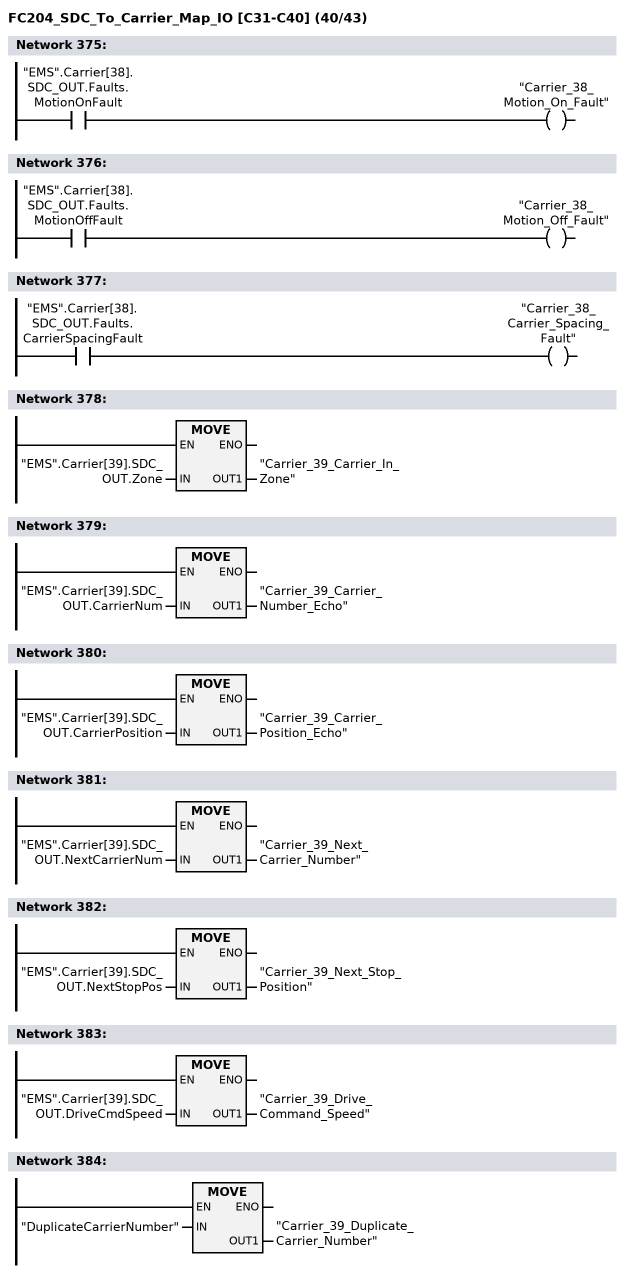
   RUNG wire#powerrail
      Contact( "EMS".Carrier[38].SDC_OUT.Faults.MotionOnFault )
      Coil( "Carrier_38_Motion_On_Fault" )
   END_RUNG
   // the same network as SCL:
   "Carrier_38_Motion_On_Fault" := "EMS".Carrier[38].SDC_OUT.Faults.MotionOnFault;
END_REGION

REGION Network 376
   RUNG wire#powerrail
      Contact( "EMS".Carrier[38].SDC_OUT.Faults.MotionOffFault )
      Coil( "Carrier_38_Motion_Off_Fault" )
   END_RUNG
   // the same network as SCL:
   "Carrier_38_Motion_Off_Fault" := "EMS".Carrier[38].SDC_OUT.Faults.MotionOffFault;
END_REGION

REGION Network 377
   RUNG wire#powerrail
      Contact( "EMS".Carrier[38].SDC_OUT.Faults.CarrierSpacingFault )
      Coil( "Carrier_38_Carrier_Spacing_Fault" )
   END_RUNG
   // the same network as SCL:
   "Carrier_38_Carrier_Spacing_Fault" := "EMS".Carrier[38].SDC_OUT.Faults.CarrierSpacingFault;
END_REGION

REGION Network 378
   RUNG wire#powerrail
      Move(in := "EMS".Carrier[39].SDC_OUT.Zone, out1 => "Carrier_39_Carrier_In_Zone")
   END_RUNG
   // the same network as SCL:
   "Carrier_39_Carrier_In_Zone" := "EMS".Carrier[39].SDC_OUT.Zone;
END_REGION

REGION Network 379
   RUNG wire#powerrail
      Move(in := "EMS".Carrier[39].SDC_OUT.CarrierNum, out1 => "Carrier_39_Carrier_Number_Echo")
   END_RUNG
   // the same network as SCL:
   "Carrier_39_Carrier_Number_Echo" := "EMS".Carrier[39].SDC_OUT.CarrierNum;
END_REGION

REGION Network 380
   RUNG wire#powerrail
      Move(in := "EMS".Carrier[39].SDC_OUT.CarrierPosition, out1 => "Carrier_39_Carrier_Position_Echo")
   END_RUNG
   // the same network as SCL:
   "Carrier_39_Carrier_Position_Echo" := "EMS".Carrier[39].SDC_OUT.CarrierPosition;
END_REGION

REGION Network 381
   RUNG wire#powerrail
      Move(in := "EMS".Carrier[39].SDC_OUT.NextCarrierNum, out1 => "Carrier_39_Next_Carrier_Number")
   END_RUNG
   // the same network as SCL:
   "Carrier_39_Next_Carrier_Number" := "EMS".Carrier[39].SDC_OUT.NextCarrierNum;
END_REGION

REGION Network 382
   RUNG wire#powerrail
      Move(in := "EMS".Carrier[39].SDC_OUT.NextStopPos, out1 => "Carrier_39_Next_Stop_Position")
   END_RUNG
   // the same network as SCL:
   "Carrier_39_Next_Stop_Position" := "EMS".Carrier[39].SDC_OUT.NextStopPos;
END_REGION

REGION Network 383
   RUNG wire#powerrail
      Move(in := "EMS".Carrier[39].SDC_OUT.DriveCmdSpeed, out1 => "Carrier_39_Drive_Command_Speed")
   END_RUNG
   // the same network as SCL:
   "Carrier_39_Drive_Command_Speed" := "EMS".Carrier[39].SDC_OUT.DriveCmdSpeed;
END_REGION

REGION Network 384
   RUNG wire#powerrail
      Move(in := "DuplicateCarrierNumber", out1 => "Carrier_39_Duplicate_Carrier_Number")
   END_RUNG
   // the same network as SCL:
   "Carrier_39_Duplicate_Carrier_Number" := "DuplicateCarrierNumber";
END_REGION

REGION Network 385
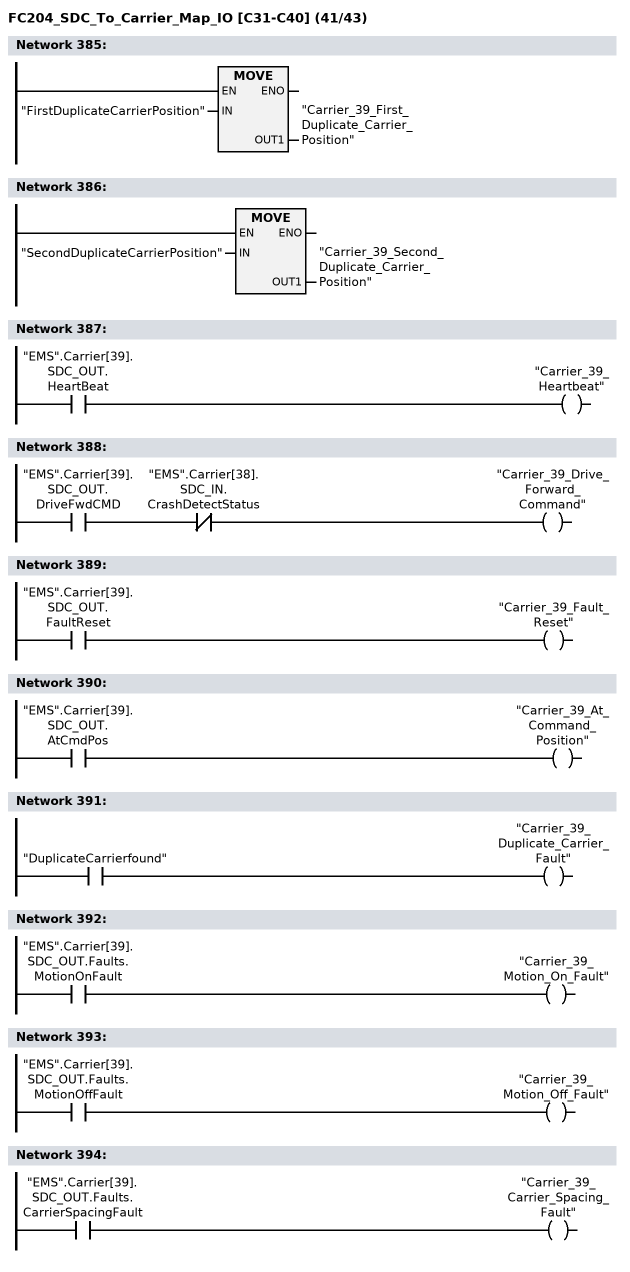
   RUNG wire#powerrail
      Move(in := "FirstDuplicateCarrierPosition", out1 => "Carrier_39_First_Duplicate_Carrier_Position")
   END_RUNG
   // the same network as SCL:
   "Carrier_39_First_Duplicate_Carrier_Position" := "FirstDuplicateCarrierPosition";
END_REGION

REGION Network 386
   RUNG wire#powerrail
      Move(in := "SecondDuplicateCarrierPosition", out1 => "Carrier_39_Second_Duplicate_Carrier_Position")
   END_RUNG
   // the same network as SCL:
   "Carrier_39_Second_Duplicate_Carrier_Position" := "SecondDuplicateCarrierPosition";
END_REGION

REGION Network 387
   RUNG wire#powerrail
      Contact( "EMS".Carrier[39].SDC_OUT.HeartBeat )
      Coil( "Carrier_39_Heartbeat" )
   END_RUNG
   // the same network as SCL:
   "Carrier_39_Heartbeat" := "EMS".Carrier[39].SDC_OUT.HeartBeat;
END_REGION

REGION Network 388
   RUNG wire#powerrail
      Contact( "EMS".Carrier[39].SDC_OUT.DriveFwdCMD )
      I_Contact( "EMS".Carrier[38].SDC_IN.CrashDetectStatus )
      Coil( "Carrier_39_Drive_Forward_Command" )
   END_RUNG
   // the same network as SCL:
   "Carrier_39_Drive_Forward_Command" := "EMS".Carrier[39].SDC_OUT.DriveFwdCMD AND NOT "EMS".Carrier[38].SDC_IN.CrashDetectStatus;
END_REGION

REGION Network 389
   RUNG wire#powerrail
      Contact( "EMS".Carrier[39].SDC_OUT.FaultReset )
      Coil( "Carrier_39_Fault_Reset" )
   END_RUNG
   // the same network as SCL:
   "Carrier_39_Fault_Reset" := "EMS".Carrier[39].SDC_OUT.FaultReset;
END_REGION

REGION Network 390
   RUNG wire#powerrail
      Contact( "EMS".Carrier[39].SDC_OUT.AtCmdPos )
      Coil( "Carrier_39_At_Command_Position" )
   END_RUNG
   // the same network as SCL:
   "Carrier_39_At_Command_Position" := "EMS".Carrier[39].SDC_OUT.AtCmdPos;
END_REGION

REGION Network 391
   RUNG wire#powerrail
      Contact( "DuplicateCarrierfound" )
      Coil( "Carrier_39_Duplicate_Carrier_Fault" )
   END_RUNG
   // the same network as SCL:
   "Carrier_39_Duplicate_Carrier_Fault" := "DuplicateCarrierfound";
END_REGION

REGION Network 392
   RUNG wire#powerrail
      Contact( "EMS".Carrier[39].SDC_OUT.Faults.MotionOnFault )
      Coil( "Carrier_39_Motion_On_Fault" )
   END_RUNG
   // the same network as SCL:
   "Carrier_39_Motion_On_Fault" := "EMS".Carrier[39].SDC_OUT.Faults.MotionOnFault;
END_REGION

REGION Network 393
   RUNG wire#powerrail
      Contact( "EMS".Carrier[39].SDC_OUT.Faults.MotionOffFault )
      Coil( "Carrier_39_Motion_Off_Fault" )
   END_RUNG
   // the same network as SCL:
   "Carrier_39_Motion_Off_Fault" := "EMS".Carrier[39].SDC_OUT.Faults.MotionOffFault;
END_REGION

REGION Network 394
   RUNG wire#powerrail
      Contact( "EMS".Carrier[39].SDC_OUT.Faults.CarrierSpacingFault )
      Coil( "Carrier_39_Carrier_Spacing_Fault" )
   END_RUNG
   // the same network as SCL:
   "Carrier_39_Carrier_Spacing_Fault" := "EMS".Carrier[39].SDC_OUT.Faults.CarrierSpacingFault;
END_REGION

REGION Network 395
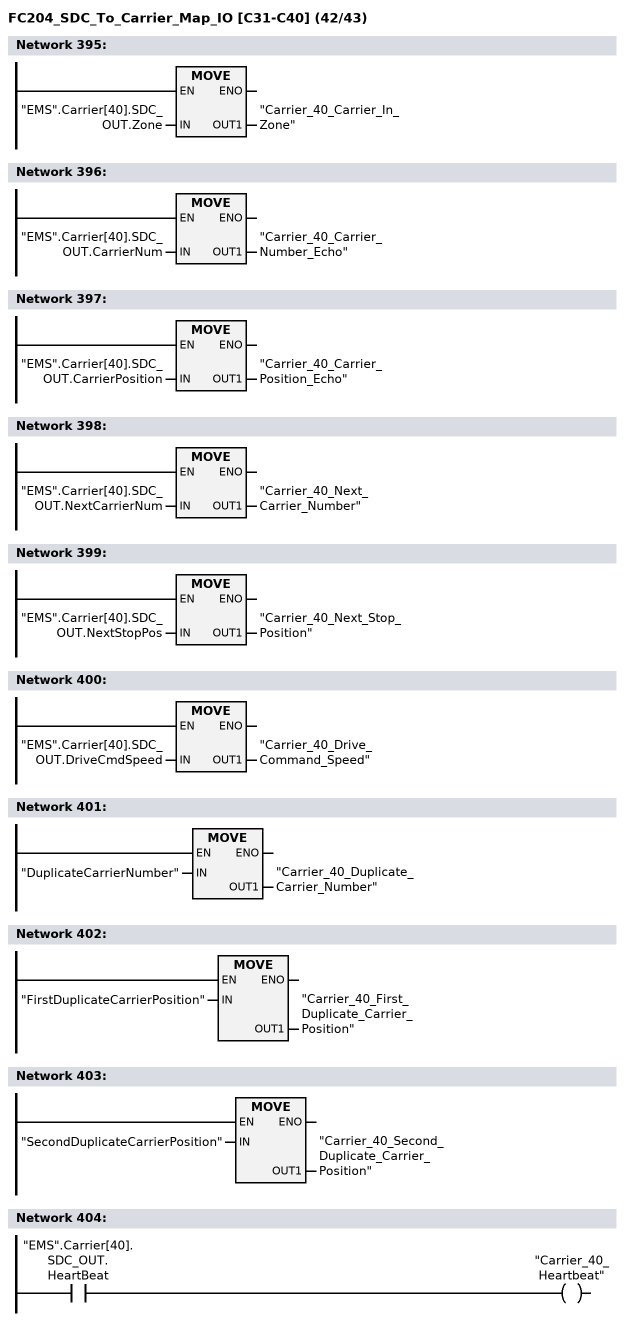
   RUNG wire#powerrail
      Move(in := "EMS".Carrier[40].SDC_OUT.Zone, out1 => "Carrier_40_Carrier_In_Zone")
   END_RUNG
   // the same network as SCL:
   "Carrier_40_Carrier_In_Zone" := "EMS".Carrier[40].SDC_OUT.Zone;
END_REGION

REGION Network 396
   RUNG wire#powerrail
      Move(in := "EMS".Carrier[40].SDC_OUT.CarrierNum, out1 => "Carrier_40_Carrier_Number_Echo")
   END_RUNG
   // the same network as SCL:
   "Carrier_40_Carrier_Number_Echo" := "EMS".Carrier[40].SDC_OUT.CarrierNum;
END_REGION

REGION Network 397
   RUNG wire#powerrail
      Move(in := "EMS".Carrier[40].SDC_OUT.CarrierPosition, out1 => "Carrier_40_Carrier_Position_Echo")
   END_RUNG
   // the same network as SCL:
   "Carrier_40_Carrier_Position_Echo" := "EMS".Carrier[40].SDC_OUT.CarrierPosition;
END_REGION

REGION Network 398
   RUNG wire#powerrail
      Move(in := "EMS".Carrier[40].SDC_OUT.NextCarrierNum, out1 => "Carrier_40_Next_Carrier_Number")
   END_RUNG
   // the same network as SCL:
   "Carrier_40_Next_Carrier_Number" := "EMS".Carrier[40].SDC_OUT.NextCarrierNum;
END_REGION

REGION Network 399
   RUNG wire#powerrail
      Move(in := "EMS".Carrier[40].SDC_OUT.NextStopPos, out1 => "Carrier_40_Next_Stop_Position")
   END_RUNG
   // the same network as SCL:
   "Carrier_40_Next_Stop_Position" := "EMS".Carrier[40].SDC_OUT.NextStopPos;
END_REGION

REGION Network 400
   RUNG wire#powerrail
      Move(in := "EMS".Carrier[40].SDC_OUT.DriveCmdSpeed, out1 => "Carrier_40_Drive_Command_Speed")
   END_RUNG
   // the same network as SCL:
   "Carrier_40_Drive_Command_Speed" := "EMS".Carrier[40].SDC_OUT.DriveCmdSpeed;
END_REGION

REGION Network 401
   RUNG wire#powerrail
      Move(in := "DuplicateCarrierNumber", out1 => "Carrier_40_Duplicate_Carrier_Number")
   END_RUNG
   // the same network as SCL:
   "Carrier_40_Duplicate_Carrier_Number" := "DuplicateCarrierNumber";
END_REGION

REGION Network 402
   RUNG wire#powerrail
      Move(in := "FirstDuplicateCarrierPosition", out1 => "Carrier_40_First_Duplicate_Carrier_Position")
   END_RUNG
   // the same network as SCL:
   "Carrier_40_First_Duplicate_Carrier_Position" := "FirstDuplicateCarrierPosition";
END_REGION

REGION Network 403
   RUNG wire#powerrail
      Move(in := "SecondDuplicateCarrierPosition", out1 => "Carrier_40_Second_Duplicate_Carrier_Position")
   END_RUNG
   // the same network as SCL:
   "Carrier_40_Second_Duplicate_Carrier_Position" := "SecondDuplicateCarrierPosition";
END_REGION

REGION Network 404
   RUNG wire#powerrail
      Contact( "EMS".Carrier[40].SDC_OUT.HeartBeat )
      Coil( "Carrier_40_Heartbeat" )
   END_RUNG
   // the same network as SCL:
   "Carrier_40_Heartbeat" := "EMS".Carrier[40].SDC_OUT.HeartBeat;
END_REGION

REGION Network 405
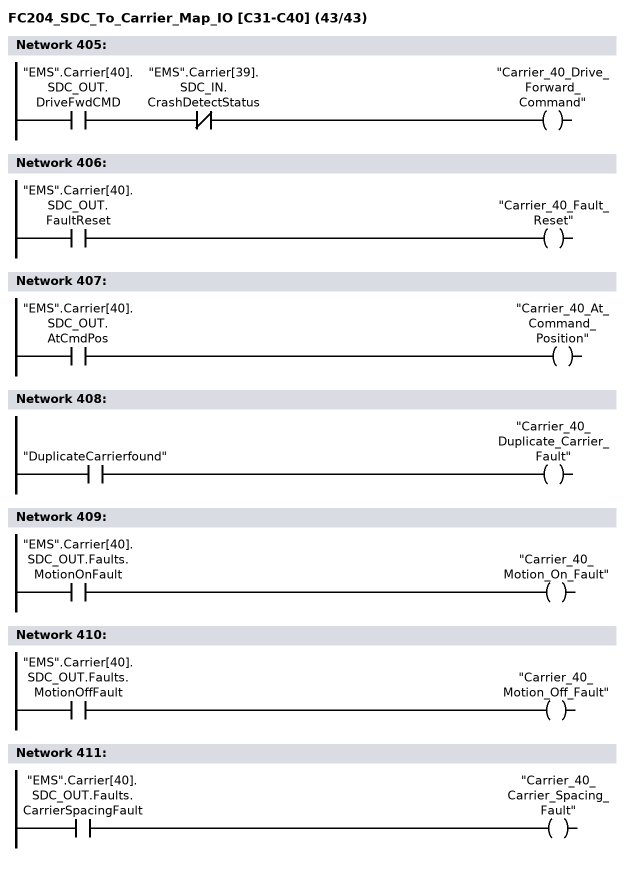
   RUNG wire#powerrail
      Contact( "EMS".Carrier[40].SDC_OUT.DriveFwdCMD )
      I_Contact( "EMS".Carrier[39].SDC_IN.CrashDetectStatus )
      Coil( "Carrier_40_Drive_Forward_Command" )
   END_RUNG
   // the same network as SCL:
   "Carrier_40_Drive_Forward_Command" := "EMS".Carrier[40].SDC_OUT.DriveFwdCMD AND NOT "EMS".Carrier[39].SDC_IN.CrashDetectStatus;
END_REGION

REGION Network 406
   RUNG wire#powerrail
      Contact( "EMS".Carrier[40].SDC_OUT.FaultReset )
      Coil( "Carrier_40_Fault_Reset" )
   END_RUNG
   // the same network as SCL:
   "Carrier_40_Fault_Reset" := "EMS".Carrier[40].SDC_OUT.FaultReset;
END_REGION

REGION Network 407
   RUNG wire#powerrail
      Contact( "EMS".Carrier[40].SDC_OUT.AtCmdPos )
      Coil( "Carrier_40_At_Command_Position" )
   END_RUNG
   // the same network as SCL:
   "Carrier_40_At_Command_Position" := "EMS".Carrier[40].SDC_OUT.AtCmdPos;
END_REGION

REGION Network 408
   RUNG wire#powerrail
      Contact( "DuplicateCarrierfound" )
      Coil( "Carrier_40_Duplicate_Carrier_Fault" )
   END_RUNG
   // the same network as SCL:
   "Carrier_40_Duplicate_Carrier_Fault" := "DuplicateCarrierfound";
END_REGION

REGION Network 409
   RUNG wire#powerrail
      Contact( "EMS".Carrier[40].SDC_OUT.Faults.MotionOnFault )
      Coil( "Carrier_40_Motion_On_Fault" )
   END_RUNG
   // the same network as SCL:
   "Carrier_40_Motion_On_Fault" := "EMS".Carrier[40].SDC_OUT.Faults.MotionOnFault;
END_REGION

REGION Network 410
   RUNG wire#powerrail
      Contact( "EMS".Carrier[40].SDC_OUT.Faults.MotionOffFault )
      Coil( "Carrier_40_Motion_Off_Fault" )
   END_RUNG
   // the same network as SCL:
   "Carrier_40_Motion_Off_Fault" := "EMS".Carrier[40].SDC_OUT.Faults.MotionOffFault;
END_REGION

REGION Network 411
   RUNG wire#powerrail
      Contact( "EMS".Carrier[40].SDC_OUT.Faults.CarrierSpacingFault )
      Coil( "Carrier_40_Carrier_Spacing_Fault" )
   END_RUNG
   // the same network as SCL:
   "Carrier_40_Carrier_Spacing_Fault" := "EMS".Carrier[40].SDC_OUT.Faults.CarrierSpacingFault;
END_REGION
END_FUNCTION

FUNCTION "FC205_SDC_To_Carrier_Map_IO [C41-C50]" : Void   // FC205, LAD
{ S7_Optimized_Access := 'TRUE' }
VERSION : 0.1
BEGIN

REGION Network 1
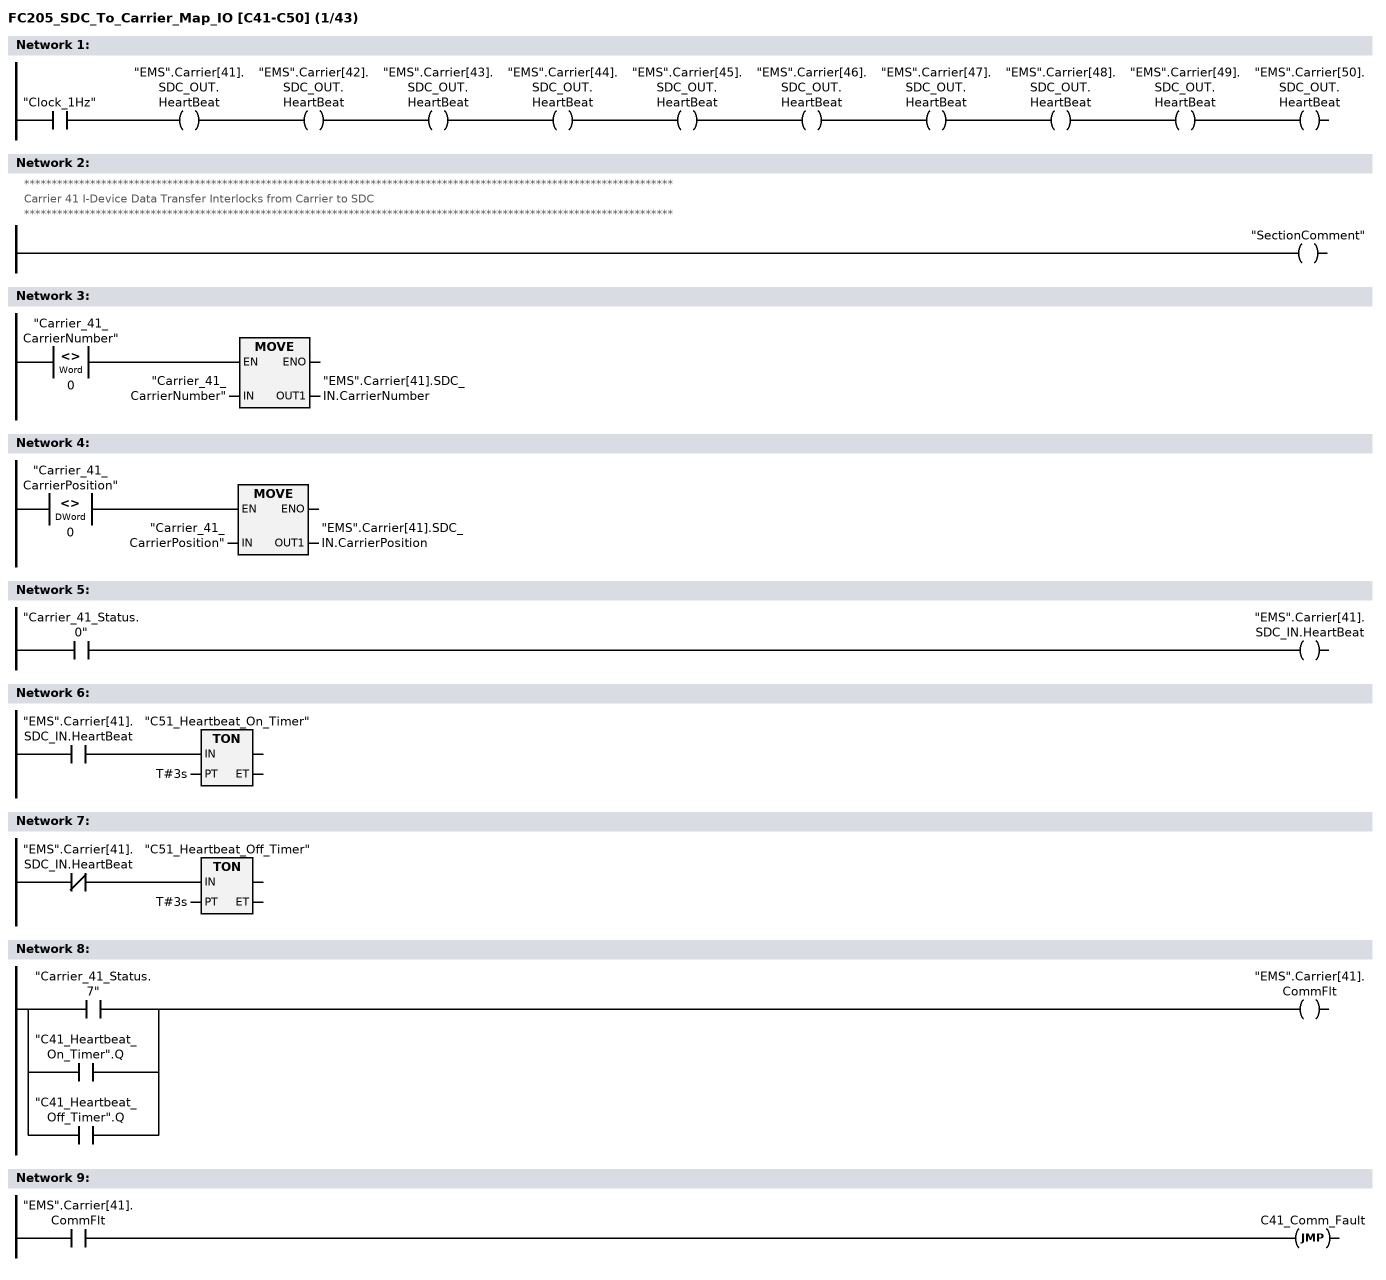
   RUNG wire#powerrail
      Contact( "Clock_1Hz" )
      Coil( "EMS".Carrier[41].SDC_OUT.HeartBeat )
      Coil( "EMS".Carrier[42].SDC_OUT.HeartBeat )
      Coil( "EMS".Carrier[43].SDC_OUT.HeartBeat )
      Coil( "EMS".Carrier[44].SDC_OUT.HeartBeat )
      Coil( "EMS".Carrier[45].SDC_OUT.HeartBeat )
      Coil( "EMS".Carrier[46].SDC_OUT.HeartBeat )
      Coil( "EMS".Carrier[47].SDC_OUT.HeartBeat )
      Coil( "EMS".Carrier[48].SDC_OUT.HeartBeat )
      Coil( "EMS".Carrier[49].SDC_OUT.HeartBeat )
      Coil( "EMS".Carrier[50].SDC_OUT.HeartBeat )
   END_RUNG
   // the same network as SCL:
   "EMS".Carrier[41].SDC_OUT.HeartBeat := "Clock_1Hz";
   "EMS".Carrier[42].SDC_OUT.HeartBeat := "Clock_1Hz";
   "EMS".Carrier[43].SDC_OUT.HeartBeat := "Clock_1Hz";
   "EMS".Carrier[44].SDC_OUT.HeartBeat := "Clock_1Hz";
   "EMS".Carrier[45].SDC_OUT.HeartBeat := "Clock_1Hz";
   "EMS".Carrier[46].SDC_OUT.HeartBeat := "Clock_1Hz";
   "EMS".Carrier[47].SDC_OUT.HeartBeat := "Clock_1Hz";
   "EMS".Carrier[48].SDC_OUT.HeartBeat := "Clock_1Hz";
   "EMS".Carrier[49].SDC_OUT.HeartBeat := "Clock_1Hz";
   "EMS".Carrier[50].SDC_OUT.HeartBeat := "Clock_1Hz";
END_REGION

REGION Network 2
   // **********************************************************************************************************************
   // 
   // Carrier 41 I-Device Data Transfer Interlocks from Carrier to SDC
   // 
   // **********************************************************************************************************************
   RUNG wire#powerrail
      Coil( "SectionComment" )
   END_RUNG
   // the same network as SCL:
   "SectionComment" := TRUE;
END_REGION

REGION Network 3
   RUNG wire#powerrail
      { S7_Templates := "SrcType := Word" } NE_Contact(in1 := "Carrier_41_CarrierNumber", in2 := 0)
      Move(in := "Carrier_41_CarrierNumber", out1 => "EMS".Carrier[41].SDC_IN.CarrierNumber)
   END_RUNG
   // the same network as SCL:
   IF "Carrier_41_CarrierNumber" <> 0 THEN
       "EMS".Carrier[41].SDC_IN.CarrierNumber := "Carrier_41_CarrierNumber";
   END_IF;
END_REGION

REGION Network 4
   RUNG wire#powerrail
      { S7_Templates := "SrcType := DWord" } NE_Contact(in1 := "Carrier_41_CarrierPosition", in2 := 0)
      Move(in := "Carrier_41_CarrierPosition", out1 => "EMS".Carrier[41].SDC_IN.CarrierPosition)
   END_RUNG
   // the same network as SCL:
   IF "Carrier_41_CarrierPosition" <> 0 THEN
       "EMS".Carrier[41].SDC_IN.CarrierPosition := "Carrier_41_CarrierPosition";
   END_IF;
END_REGION

REGION Network 5
   RUNG wire#powerrail
      Contact( "Carrier_41_Status.0" )
      Coil( "EMS".Carrier[41].SDC_IN.HeartBeat )
   END_RUNG
   // the same network as SCL:
   "EMS".Carrier[41].SDC_IN.HeartBeat := "Carrier_41_Status.0";
END_REGION

REGION Network 6
   "C51_Heartbeat_On_Timer".TON(IN := "EMS".Carrier[41].SDC_IN.HeartBeat, PT := T#3s);
END_REGION

REGION Network 7
   "C51_Heartbeat_Off_Timer".TON(IN := NOT "EMS".Carrier[41].SDC_IN.HeartBeat, PT := T#3s);
END_REGION

REGION Network 8
   RUNG wire#powerrail
      Contact( "Carrier_41_Status.7" )
      wire#w1
      Coil( "EMS".Carrier[41].CommFlt )
   END_RUNG
   RUNG wire#powerrail
      Contact( "C41_Heartbeat_On_Timer".Q )
   END_RUNG wire#w1
   RUNG wire#powerrail
      Contact( "C41_Heartbeat_Off_Timer".Q )
   END_RUNG wire#w1
   // the same network as SCL:
   "EMS".Carrier[41].CommFlt := "Carrier_41_Status.7" OR "C41_Heartbeat_On_Timer".Q OR "C41_Heartbeat_Off_Timer".Q;
END_REGION

REGION Network 9
   RUNG wire#powerrail
      Contact( "EMS".Carrier[41].CommFlt )
      JumpCoil( C41_Comm_Fault )
   END_RUNG
   // the same network as SCL:
   IF "EMS".Carrier[41].CommFlt THEN GOTO C41_Comm_Fault; END_IF;
END_REGION

REGION Network 10
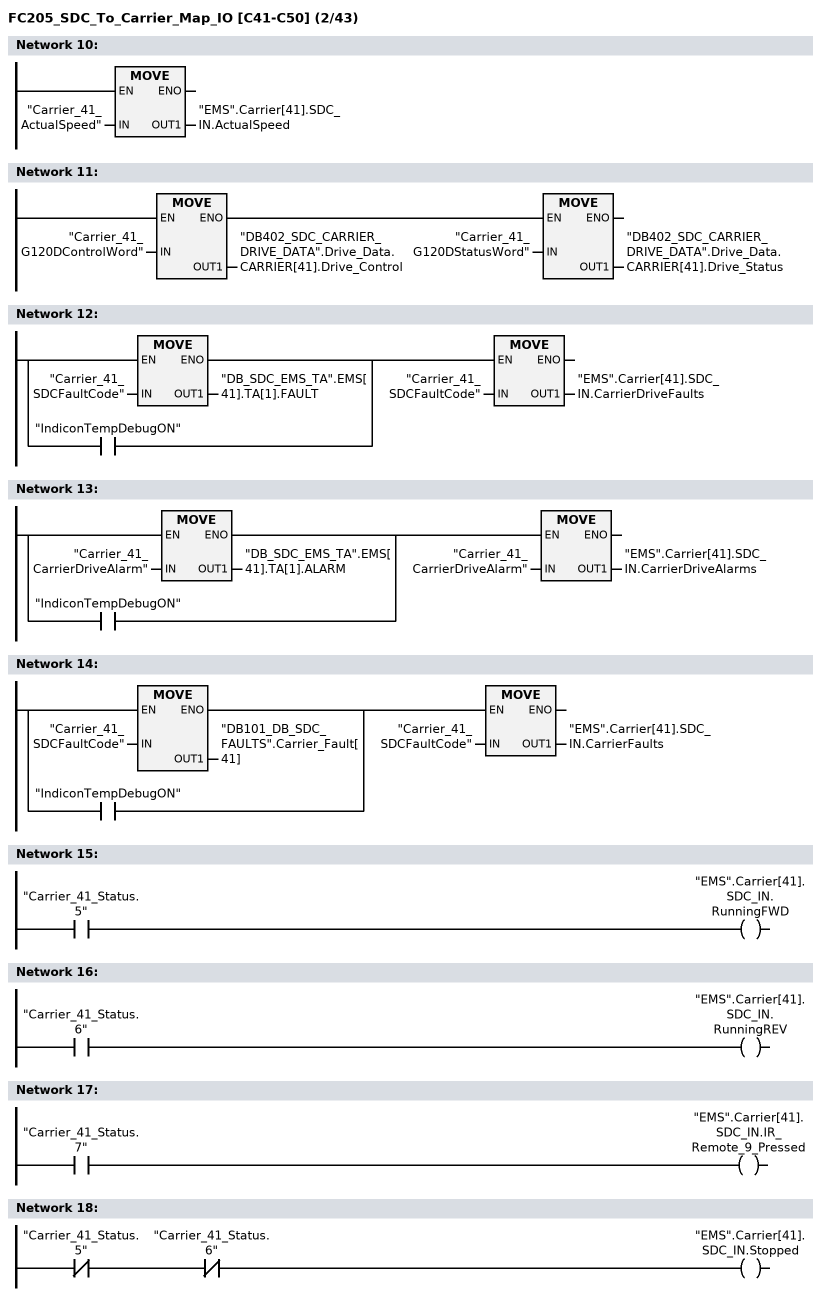
   RUNG wire#powerrail
      Move(in := "Carrier_41_ActualSpeed", out1 => "EMS".Carrier[41].SDC_IN.ActualSpeed)
   END_RUNG
   // the same network as SCL:
   "EMS".Carrier[41].SDC_IN.ActualSpeed := "Carrier_41_ActualSpeed";
END_REGION

REGION Network 11
   RUNG wire#powerrail
      Move(in := "Carrier_41_G120DControlWord", out1 => "DB402_SDC_CARRIER_DRIVE_DATA".Drive_Data.CARRIER[41].Drive_Control)
      Move(in := "Carrier_41_G120DStatusWord", out1 => "DB402_SDC_CARRIER_DRIVE_DATA".Drive_Data.CARRIER[41].Drive_Status)
   END_RUNG
   // the same network as SCL:
   "DB402_SDC_CARRIER_DRIVE_DATA".Drive_Data.CARRIER[41].Drive_Control := "Carrier_41_G120DControlWord";
   "DB402_SDC_CARRIER_DRIVE_DATA".Drive_Data.CARRIER[41].Drive_Status := "Carrier_41_G120DStatusWord";
END_REGION

REGION Network 12
   RUNG wire#powerrail
      Move(in := "Carrier_41_SDCFaultCode", out1 => "DB_SDC_EMS_TA".EMS[41].TA[1].FAULT)
      wire#w1
      Move(in := "Carrier_41_SDCFaultCode", out1 => "EMS".Carrier[41].SDC_IN.CarrierDriveFaults)
   END_RUNG
   RUNG wire#powerrail
      Contact( "IndiconTempDebugON" )
   END_RUNG wire#w1
   // the same network as SCL:
   "DB_SDC_EMS_TA".EMS[41].TA[1].FAULT := "Carrier_41_SDCFaultCode";
   IF TRUE OR "IndiconTempDebugON" THEN
       "EMS".Carrier[41].SDC_IN.CarrierDriveFaults := "Carrier_41_SDCFaultCode";
   END_IF;
END_REGION

REGION Network 13
   RUNG wire#powerrail
      Move(in := "Carrier_41_CarrierDriveAlarm", out1 => "DB_SDC_EMS_TA".EMS[41].TA[1].ALARM)
      wire#w1
      Move(in := "Carrier_41_CarrierDriveAlarm", out1 => "EMS".Carrier[41].SDC_IN.CarrierDriveAlarms)
   END_RUNG
   RUNG wire#powerrail
      Contact( "IndiconTempDebugON" )
   END_RUNG wire#w1
   // the same network as SCL:
   "DB_SDC_EMS_TA".EMS[41].TA[1].ALARM := "Carrier_41_CarrierDriveAlarm";
   IF TRUE OR "IndiconTempDebugON" THEN
       "EMS".Carrier[41].SDC_IN.CarrierDriveAlarms := "Carrier_41_CarrierDriveAlarm";
   END_IF;
END_REGION

REGION Network 14
   RUNG wire#powerrail
      Move(in := "Carrier_41_SDCFaultCode", out1 => "DB101_DB_SDC_FAULTS".Carrier_Fault[41])
      wire#w1
      Move(in := "Carrier_41_SDCFaultCode", out1 => "EMS".Carrier[41].SDC_IN.CarrierFaults)
   END_RUNG
   RUNG wire#powerrail
      Contact( "IndiconTempDebugON" )
   END_RUNG wire#w1
   // the same network as SCL:
   "DB101_DB_SDC_FAULTS".Carrier_Fault[41] := "Carrier_41_SDCFaultCode";
   IF TRUE OR "IndiconTempDebugON" THEN
       "EMS".Carrier[41].SDC_IN.CarrierFaults := "Carrier_41_SDCFaultCode";
   END_IF;
END_REGION

REGION Network 15
   RUNG wire#powerrail
      Contact( "Carrier_41_Status.5" )
      Coil( "EMS".Carrier[41].SDC_IN.RunningFWD )
   END_RUNG
   // the same network as SCL:
   "EMS".Carrier[41].SDC_IN.RunningFWD := "Carrier_41_Status.5";
END_REGION

REGION Network 16
   RUNG wire#powerrail
      Contact( "Carrier_41_Status.6" )
      Coil( "EMS".Carrier[41].SDC_IN.RunningREV )
   END_RUNG
   // the same network as SCL:
   "EMS".Carrier[41].SDC_IN.RunningREV := "Carrier_41_Status.6";
END_REGION

REGION Network 17
   RUNG wire#powerrail
      Contact( "Carrier_41_Status.7" )
      Coil( "EMS".Carrier[41].SDC_IN.IR_Remote_9_Pressed )
   END_RUNG
   // the same network as SCL:
   "EMS".Carrier[41].SDC_IN.IR_Remote_9_Pressed := "Carrier_41_Status.7";
END_REGION

REGION Network 18
   RUNG wire#powerrail
      I_Contact( "Carrier_41_Status.5" )
      I_Contact( "Carrier_41_Status.6" )
      Coil( "EMS".Carrier[41].SDC_IN.Stopped )
   END_RUNG
   // the same network as SCL:
   "EMS".Carrier[41].SDC_IN.Stopped := NOT "Carrier_41_Status.5" AND NOT "Carrier_41_Status.6";
END_REGION

REGION Network 19
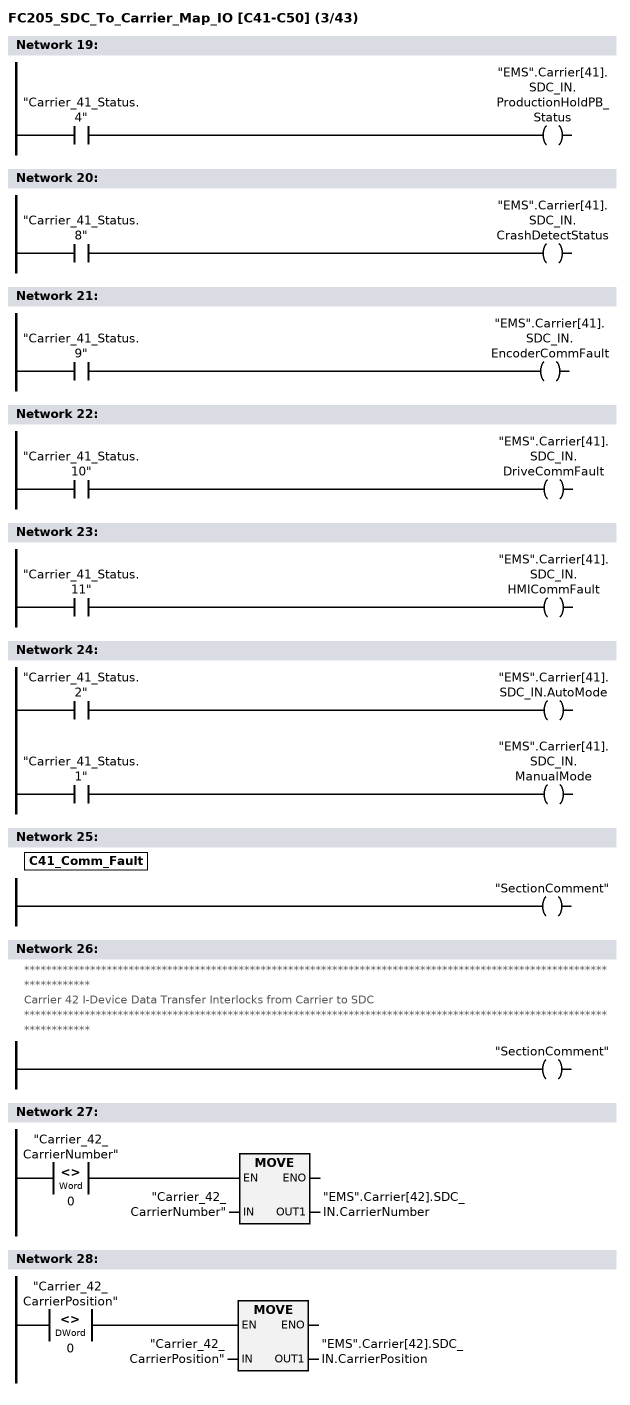
   RUNG wire#powerrail
      Contact( "Carrier_41_Status.4" )
      Coil( "EMS".Carrier[41].SDC_IN.ProductionHoldPB_Status )
   END_RUNG
   // the same network as SCL:
   "EMS".Carrier[41].SDC_IN.ProductionHoldPB_Status := "Carrier_41_Status.4";
END_REGION

REGION Network 20
   RUNG wire#powerrail
      Contact( "Carrier_41_Status.8" )
      Coil( "EMS".Carrier[41].SDC_IN.CrashDetectStatus )
   END_RUNG
   // the same network as SCL:
   "EMS".Carrier[41].SDC_IN.CrashDetectStatus := "Carrier_41_Status.8";
END_REGION

REGION Network 21
   RUNG wire#powerrail
      Contact( "Carrier_41_Status.9" )
      Coil( "EMS".Carrier[41].SDC_IN.EncoderCommFault )
   END_RUNG
   // the same network as SCL:
   "EMS".Carrier[41].SDC_IN.EncoderCommFault := "Carrier_41_Status.9";
END_REGION

REGION Network 22
   RUNG wire#powerrail
      Contact( "Carrier_41_Status.10" )
      Coil( "EMS".Carrier[41].SDC_IN.DriveCommFault )
   END_RUNG
   // the same network as SCL:
   "EMS".Carrier[41].SDC_IN.DriveCommFault := "Carrier_41_Status.10";
END_REGION

REGION Network 23
   RUNG wire#powerrail
      Contact( "Carrier_41_Status.11" )
      Coil( "EMS".Carrier[41].SDC_IN.HMICommFault )
   END_RUNG
   // the same network as SCL:
   "EMS".Carrier[41].SDC_IN.HMICommFault := "Carrier_41_Status.11";
END_REGION

REGION Network 24
   RUNG wire#powerrail
      Contact( "Carrier_41_Status.2" )
      Coil( "EMS".Carrier[41].SDC_IN.AutoMode )
   END_RUNG
   RUNG wire#powerrail
      Contact( "Carrier_41_Status.1" )
      Coil( "EMS".Carrier[41].SDC_IN.ManualMode )
   END_RUNG
   // the same network as SCL:
   "EMS".Carrier[41].SDC_IN.AutoMode := "Carrier_41_Status.2";
   "EMS".Carrier[41].SDC_IN.ManualMode := "Carrier_41_Status.1";
END_REGION

REGION Network 25
   Label( C41_Comm_Fault )
   RUNG wire#powerrail
      Coil( "SectionComment" )
   END_RUNG
   // the same network as SCL:
   C41_Comm_Fault:
   "SectionComment" := TRUE;
END_REGION

REGION Network 26
   // **********************************************************************************************************************
   // 
   // Carrier 42 I-Device Data Transfer Interlocks from Carrier to SDC
   // 
   // **********************************************************************************************************************
   RUNG wire#powerrail
      Coil( "SectionComment" )
   END_RUNG
   // the same network as SCL:
   "SectionComment" := TRUE;
END_REGION

REGION Network 27
   RUNG wire#powerrail
      { S7_Templates := "SrcType := Word" } NE_Contact(in1 := "Carrier_42_CarrierNumber", in2 := 0)
      Move(in := "Carrier_42_CarrierNumber", out1 => "EMS".Carrier[42].SDC_IN.CarrierNumber)
   END_RUNG
   // the same network as SCL:
   IF "Carrier_42_CarrierNumber" <> 0 THEN
       "EMS".Carrier[42].SDC_IN.CarrierNumber := "Carrier_42_CarrierNumber";
   END_IF;
END_REGION

REGION Network 28
   RUNG wire#powerrail
      { S7_Templates := "SrcType := DWord" } NE_Contact(in1 := "Carrier_42_CarrierPosition", in2 := 0)
      Move(in := "Carrier_42_CarrierPosition", out1 => "EMS".Carrier[42].SDC_IN.CarrierPosition)
   END_RUNG
   // the same network as SCL:
   IF "Carrier_42_CarrierPosition" <> 0 THEN
       "EMS".Carrier[42].SDC_IN.CarrierPosition := "Carrier_42_CarrierPosition";
   END_IF;
END_REGION

REGION Network 29
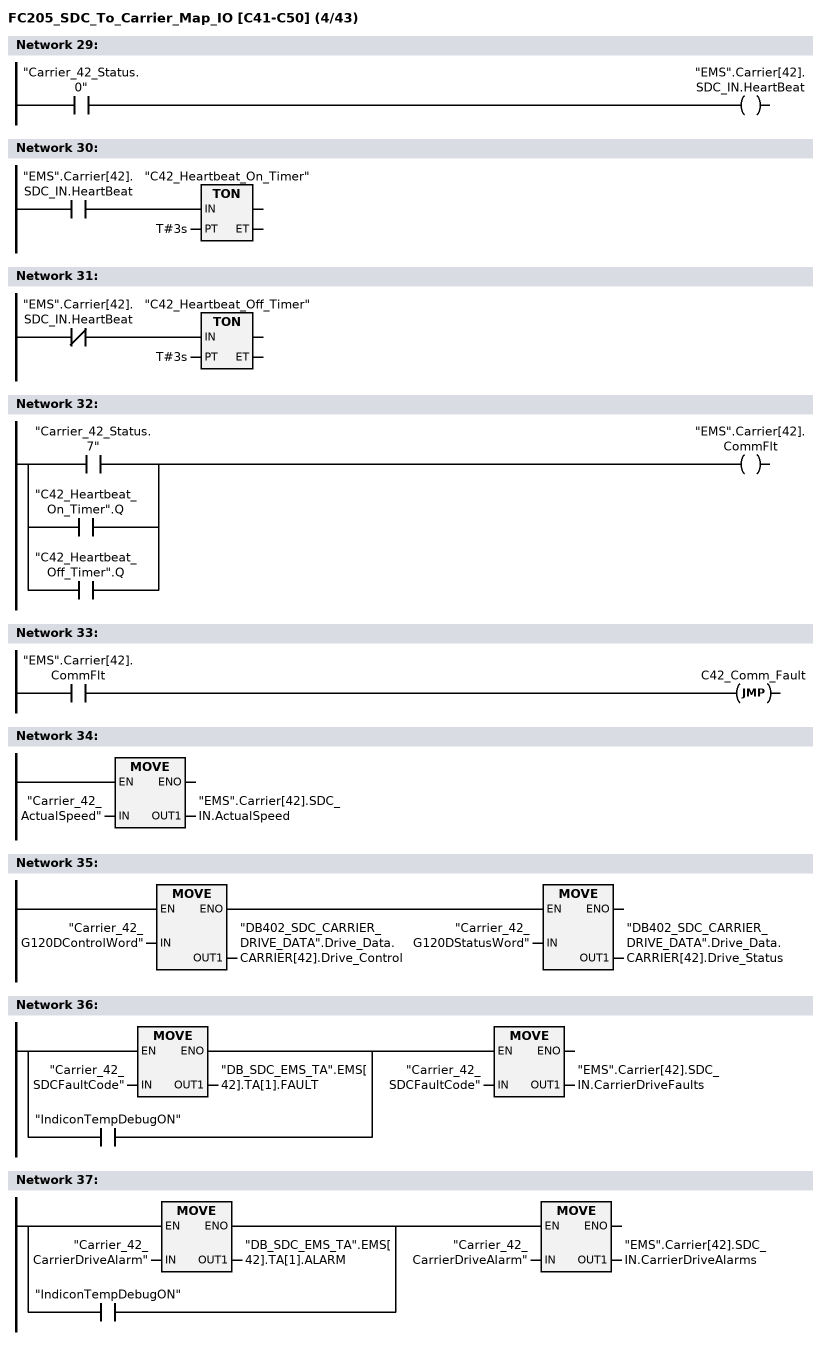
   RUNG wire#powerrail
      Contact( "Carrier_42_Status.0" )
      Coil( "EMS".Carrier[42].SDC_IN.HeartBeat )
   END_RUNG
   // the same network as SCL:
   "EMS".Carrier[42].SDC_IN.HeartBeat := "Carrier_42_Status.0";
END_REGION

REGION Network 30
   "C42_Heartbeat_On_Timer".TON(IN := "EMS".Carrier[42].SDC_IN.HeartBeat, PT := T#3s);
END_REGION

REGION Network 31
   "C42_Heartbeat_Off_Timer".TON(IN := NOT "EMS".Carrier[42].SDC_IN.HeartBeat, PT := T#3s);
END_REGION

REGION Network 32
   RUNG wire#powerrail
      Contact( "Carrier_42_Status.7" )
      wire#w1
      Coil( "EMS".Carrier[42].CommFlt )
   END_RUNG
   RUNG wire#powerrail
      Contact( "C42_Heartbeat_On_Timer".Q )
   END_RUNG wire#w1
   RUNG wire#powerrail
      Contact( "C42_Heartbeat_Off_Timer".Q )
   END_RUNG wire#w1
   // the same network as SCL:
   "EMS".Carrier[42].CommFlt := "Carrier_42_Status.7" OR "C42_Heartbeat_On_Timer".Q OR "C42_Heartbeat_Off_Timer".Q;
END_REGION

REGION Network 33
   RUNG wire#powerrail
      Contact( "EMS".Carrier[42].CommFlt )
      JumpCoil( C42_Comm_Fault )
   END_RUNG
   // the same network as SCL:
   IF "EMS".Carrier[42].CommFlt THEN GOTO C42_Comm_Fault; END_IF;
END_REGION

REGION Network 34
   RUNG wire#powerrail
      Move(in := "Carrier_42_ActualSpeed", out1 => "EMS".Carrier[42].SDC_IN.ActualSpeed)
   END_RUNG
   // the same network as SCL:
   "EMS".Carrier[42].SDC_IN.ActualSpeed := "Carrier_42_ActualSpeed";
END_REGION

REGION Network 35
   RUNG wire#powerrail
      Move(in := "Carrier_42_G120DControlWord", out1 => "DB402_SDC_CARRIER_DRIVE_DATA".Drive_Data.CARRIER[42].Drive_Control)
      Move(in := "Carrier_42_G120DStatusWord", out1 => "DB402_SDC_CARRIER_DRIVE_DATA".Drive_Data.CARRIER[42].Drive_Status)
   END_RUNG
   // the same network as SCL:
   "DB402_SDC_CARRIER_DRIVE_DATA".Drive_Data.CARRIER[42].Drive_Control := "Carrier_42_G120DControlWord";
   "DB402_SDC_CARRIER_DRIVE_DATA".Drive_Data.CARRIER[42].Drive_Status := "Carrier_42_G120DStatusWord";
END_REGION

REGION Network 36
   RUNG wire#powerrail
      Move(in := "Carrier_42_SDCFaultCode", out1 => "DB_SDC_EMS_TA".EMS[42].TA[1].FAULT)
      wire#w1
      Move(in := "Carrier_42_SDCFaultCode", out1 => "EMS".Carrier[42].SDC_IN.CarrierDriveFaults)
   END_RUNG
   RUNG wire#powerrail
      Contact( "IndiconTempDebugON" )
   END_RUNG wire#w1
   // the same network as SCL:
   "DB_SDC_EMS_TA".EMS[42].TA[1].FAULT := "Carrier_42_SDCFaultCode";
   IF TRUE OR "IndiconTempDebugON" THEN
       "EMS".Carrier[42].SDC_IN.CarrierDriveFaults := "Carrier_42_SDCFaultCode";
   END_IF;
END_REGION

REGION Network 37
   RUNG wire#powerrail
      Move(in := "Carrier_42_CarrierDriveAlarm", out1 => "DB_SDC_EMS_TA".EMS[42].TA[1].ALARM)
      wire#w1
      Move(in := "Carrier_42_CarrierDriveAlarm", out1 => "EMS".Carrier[42].SDC_IN.CarrierDriveAlarms)
   END_RUNG
   RUNG wire#powerrail
      Contact( "IndiconTempDebugON" )
   END_RUNG wire#w1
   // the same network as SCL:
   "DB_SDC_EMS_TA".EMS[42].TA[1].ALARM := "Carrier_42_CarrierDriveAlarm";
   IF TRUE OR "IndiconTempDebugON" THEN
       "EMS".Carrier[42].SDC_IN.CarrierDriveAlarms := "Carrier_42_CarrierDriveAlarm";
   END_IF;
END_REGION

REGION Network 38